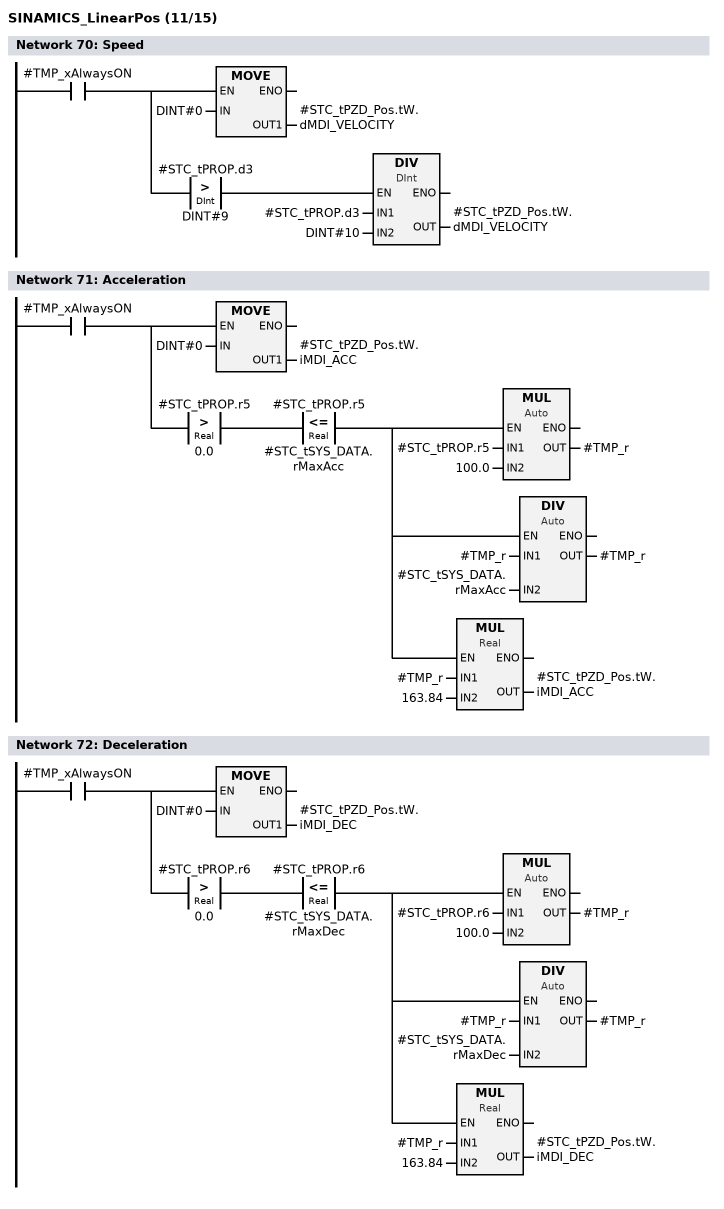
   RUNG wire#powerrail
      Contact( #TMP_xAlwaysON )
      wire#w1
      { S7_GenerateENO := "TRUE" } Move(in := DINT#0, out1 => #STC_tPZD_Pos.tW.dMDI_VELOCITY)
   END_RUNG
   RUNG wire#w1
      { S7_Templates := "SrcType := DInt" } GT_Contact(in1 := #STC_tPROP.d3, in2 := DINT#9)
      { S7_Templates := "SrcType := DInt"; S7_GenerateENO := "TRUE" } Div(in1 := #STC_tPROP.d3, in2 := DINT#10, out => #STC_tPZD_Pos.tW.dMDI_VELOCITY)
   END_RUNG
   // the same network as SCL:
   IF #TMP_xAlwaysON THEN #STC_tPZD_Pos.tW.dMDI_VELOCITY := DINT#0; END_IF;
   IF #TMP_xAlwaysON AND (#STC_tPROP.d3 > DINT#9) THEN
       #STC_tPZD_Pos.tW.dMDI_VELOCITY := #STC_tPROP.d3 / DINT#10;
   END_IF;
END_REGION

REGION Network 71: Acceleration
   RUNG wire#powerrail
      Contact( #TMP_xAlwaysON )
      wire#w1
      Move(in := DINT#0, out1 => #STC_tPZD_Pos.tW.iMDI_ACC)
   END_RUNG
   RUNG wire#w1
      { S7_Templates := "SrcType := Real" } GT_Contact(in1 := #STC_tPROP.r5, in2 := 0.0)
      { S7_Templates := "SrcType := Real" } LE_Contact(in1 := #STC_tPROP.r5, in2 := #STC_tSYS_DATA.rMaxAcc)
      wire#w2
      Mul(in1 := #STC_tPROP.r5, in2 := 100.0, out => #TMP_r)
   END_RUNG
   RUNG wire#w2
      Div(in1 := #TMP_r, in2 := #STC_tSYS_DATA.rMaxAcc, out => #TMP_r)
   END_RUNG
   RUNG wire#w2
      { S7_Templates := "SrcType := Real" } Mul(in1 := #TMP_r, in2 := 163.84, out => #STC_tPZD_Pos.tW.iMDI_ACC)
   END_RUNG
   // the same network as SCL:
   IF #TMP_xAlwaysON THEN #STC_tPZD_Pos.tW.iMDI_ACC := DINT#0; END_IF;
   IF #TMP_xAlwaysON AND (#STC_tPROP.r5 > 0.0) AND (#STC_tPROP.r5 <= #STC_tSYS_DATA.rMaxAcc) THEN
       #TMP_r := #STC_tPROP.r5 * 100.0;
       #TMP_r := #TMP_r / #STC_tSYS_DATA.rMaxAcc;
       #STC_tPZD_Pos.tW.iMDI_ACC := #TMP_r * 163.84;
   END_IF;
END_REGION

REGION Network 72: Deceleration
   RUNG wire#powerrail
      Contact( #TMP_xAlwaysON )
      wire#w1
      Move(in := DINT#0, out1 => #STC_tPZD_Pos.tW.iMDI_DEC)
   END_RUNG
   RUNG wire#w1
      { S7_Templates := "SrcType := Real" } GT_Contact(in1 := #STC_tPROP.r6, in2 := 0.0)
      { S7_Templates := "SrcType := Real" } LE_Contact(in1 := #STC_tPROP.r6, in2 := #STC_tSYS_DATA.rMaxDec)
      wire#w2
      Mul(in1 := #STC_tPROP.r6, in2 := 100.0, out => #TMP_r)
   END_RUNG
   RUNG wire#w2
      Div(in1 := #TMP_r, in2 := #STC_tSYS_DATA.rMaxDec, out => #TMP_r)
   END_RUNG
   RUNG wire#w2
      { S7_Templates := "SrcType := Real" } Mul(in1 := #TMP_r, in2 := 163.84, out => #STC_tPZD_Pos.tW.iMDI_DEC)
   END_RUNG
   // the same network as SCL:
   IF #TMP_xAlwaysON THEN #STC_tPZD_Pos.tW.iMDI_DEC := DINT#0; END_IF;
   IF #TMP_xAlwaysON AND (#STC_tPROP.r6 > 0.0) AND (#STC_tPROP.r6 <= #STC_tSYS_DATA.rMaxDec) THEN
       #TMP_r := #STC_tPROP.r6 * 100.0;
       #TMP_r := #TMP_r / #STC_tSYS_DATA.rMaxDec;
       #STC_tPZD_Pos.tW.iMDI_DEC := #TMP_r * 163.84;
   END_IF;
END_REGION

REGION Network 73: ########################_OPEN_CLOSE_LOOP_#######################
END_REGION

REGION Network 74: #####_MATCH_#####
END_REGION

REGION Network 75 (STL): Input copy
         JU    Out;

   T1:   CALL  BLKMOV
         ( SRCBLK  := #TMP_a,
           RET_VAL := #TMP_iRetVal,
           DSTBLK  := #STC_tPZD_OpCLLoop.tR
         );
END_REGION

REGION Network 76: Status signals
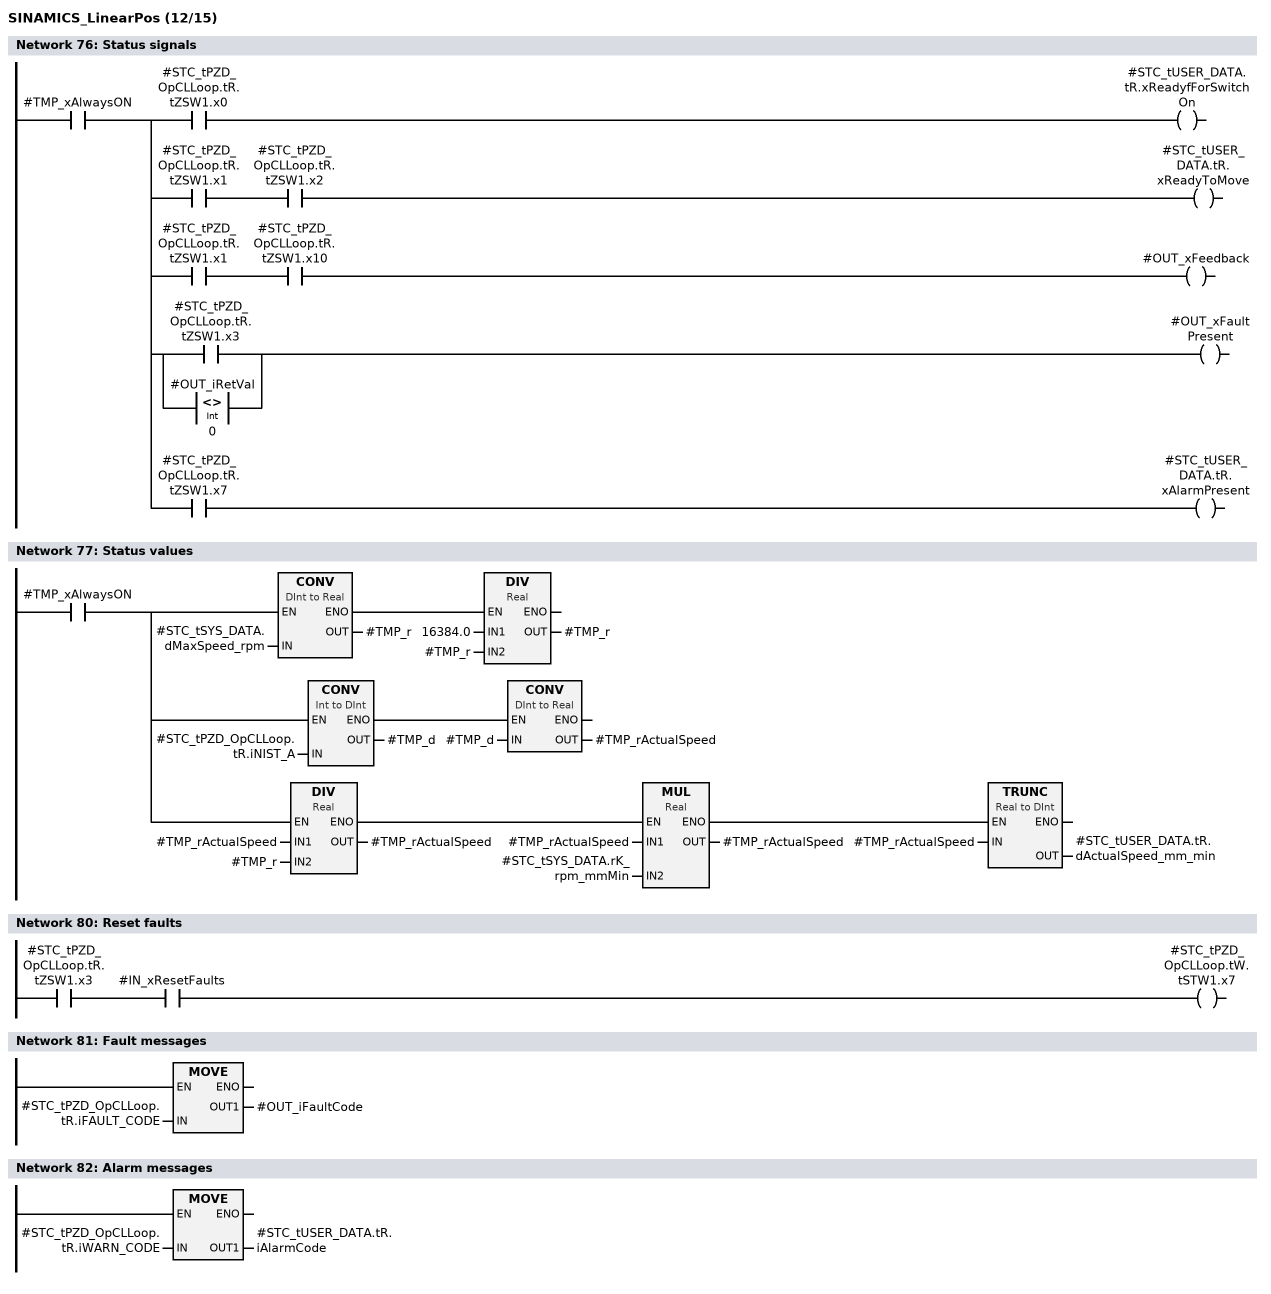
   RUNG wire#powerrail
      Contact( #TMP_xAlwaysON )
      wire#w1
      Contact( #STC_tPZD_OpCLLoop.tR.tZSW1.x0 )
      Coil( #STC_tUSER_DATA.tR.xReadyfForSwitchOn )
   END_RUNG
   RUNG wire#w1
      Contact( #STC_tPZD_OpCLLoop.tR.tZSW1.x1 )
      Contact( #STC_tPZD_OpCLLoop.tR.tZSW1.x2 )
      Coil( #STC_tUSER_DATA.tR.xReadyToMove )
   END_RUNG
   RUNG wire#w1
      Contact( #STC_tPZD_OpCLLoop.tR.tZSW1.x1 )
      Contact( #STC_tPZD_OpCLLoop.tR.tZSW1.x10 )
      Coil( #OUT_xFeedback )
   END_RUNG
   RUNG wire#w1
      Contact( #STC_tPZD_OpCLLoop.tR.tZSW1.x3 )
      wire#w2
      Coil( #OUT_xFaultPresent )
   END_RUNG
   RUNG wire#w1
      { S7_Templates := "SrcType := Int" } NE_Contact(in1 := #OUT_iRetVal, in2 := 0)
   END_RUNG wire#w2
   RUNG wire#w1
      Contact( #STC_tPZD_OpCLLoop.tR.tZSW1.x7 )
      Coil( #STC_tUSER_DATA.tR.xAlarmPresent )
   END_RUNG
   // the same network as SCL:
   #STC_tUSER_DATA.tR.xReadyfForSwitchOn := #TMP_xAlwaysON AND #STC_tPZD_OpCLLoop.tR.tZSW1.x0;
   #STC_tUSER_DATA.tR.xReadyToMove := #TMP_xAlwaysON AND #STC_tPZD_OpCLLoop.tR.tZSW1.x1 AND #STC_tPZD_OpCLLoop.tR.tZSW1.x2;
   #OUT_xFeedback := #TMP_xAlwaysON AND #STC_tPZD_OpCLLoop.tR.tZSW1.x1 AND #STC_tPZD_OpCLLoop.tR.tZSW1.x10;
   #OUT_xFaultPresent := #TMP_xAlwaysON AND (#STC_tPZD_OpCLLoop.tR.tZSW1.x3 OR (#OUT_iRetVal <> 0));
   #STC_tUSER_DATA.tR.xAlarmPresent := #TMP_xAlwaysON AND #STC_tPZD_OpCLLoop.tR.tZSW1.x7;
END_REGION

REGION Network 77: Status values
   RUNG wire#powerrail
      Contact( #TMP_xAlwaysON )
      wire#w1
      { S7_Templates := "[SrcType := DInt, DestType := Real]"; S7_GenerateENO := "TRUE" } Convert(in := #STC_tSYS_DATA.dMaxSpeed_rpm, out => #TMP_r)
      { S7_Templates := "SrcType := Real"; S7_GenerateENO := "TRUE" } Div(in1 := 16384.0, in2 := #TMP_r, out => #TMP_r)
   END_RUNG
   RUNG wire#w1
      { S7_Templates := "[SrcType := Int, DestType := DInt]"; S7_GenerateENO := "TRUE" } Convert(in := #STC_tPZD_OpCLLoop.tR.iNIST_A, out => #TMP_d)
      { S7_Templates := "[SrcType := DInt, DestType := Real]"; S7_GenerateENO := "TRUE" } Convert(in := #TMP_d, out => #TMP_rActualSpeed)
   END_RUNG
   RUNG wire#w1
      { S7_Templates := "SrcType := Real"; S7_GenerateENO := "TRUE" } Div(in1 := #TMP_rActualSpeed, in2 := #TMP_r, out => #TMP_rActualSpeed)
      { S7_Templates := "SrcType := Real"; S7_GenerateENO := "TRUE" } Mul(in1 := #TMP_rActualSpeed, in2 := #STC_tSYS_DATA.rK_rpm_mmMin, out => #TMP_rActualSpeed)
      { S7_Templates := "[SrcType := Real, DestType := DInt]"; S7_GenerateENO := "TRUE" } Trunc(in := #TMP_rActualSpeed, out => #STC_tUSER_DATA.tR.dActualSpeed_mm_min)
   END_RUNG
   // the same network as SCL:
   // ENO of a box is taken as its EN; it also drops when the box reports an error
   IF #TMP_xAlwaysON THEN
       #TMP_r := DINT_TO_REAL(#STC_tSYS_DATA.dMaxSpeed_rpm);
       #TMP_r := 16384.0 / #TMP_r;
       #TMP_d := INT_TO_DINT(#STC_tPZD_OpCLLoop.tR.iNIST_A);
       #TMP_rActualSpeed := DINT_TO_REAL(#TMP_d);
       #TMP_rActualSpeed := #TMP_rActualSpeed / #TMP_r;
       #TMP_rActualSpeed := #TMP_rActualSpeed * #STC_tSYS_DATA.rK_rpm_mmMin;
       #STC_tUSER_DATA.tR.dActualSpeed_mm_min := TRUNC(#TMP_rActualSpeed);
   END_IF;
END_REGION

REGION Network 78: #####_STATUSES_#####
END_REGION

REGION Network 79: #####_ALARMS_#####
END_REGION

REGION Network 80: Reset faults
   RUNG wire#powerrail
      Contact( #STC_tPZD_OpCLLoop.tR.tZSW1.x3 )
      Contact( #IN_xResetFaults )
      Coil( #STC_tPZD_OpCLLoop.tW.tSTW1.x7 )
   END_RUNG
   // the same network as SCL:
   #STC_tPZD_OpCLLoop.tW.tSTW1.x7 := #STC_tPZD_OpCLLoop.tR.tZSW1.x3 AND #IN_xResetFaults;
END_REGION

REGION Network 81: Fault messages
   RUNG wire#powerrail
      { S7_GenerateENO := "TRUE" } Move(in := #STC_tPZD_OpCLLoop.tR.iFAULT_CODE, out1 => #OUT_iFaultCode)
   END_RUNG
   // the same network as SCL:
   #OUT_iFaultCode := #STC_tPZD_OpCLLoop.tR.iFAULT_CODE;
END_REGION

REGION Network 82: Alarm messages
   RUNG wire#powerrail
      { S7_GenerateENO := "TRUE" } Move(in := #STC_tPZD_OpCLLoop.tR.iWARN_CODE, out1 => #STC_tUSER_DATA.tR.iAlarmCode)
   END_RUNG
   // the same network as SCL:
   #STC_tUSER_DATA.tR.iAlarmCode := #STC_tPZD_OpCLLoop.tR.iWARN_CODE;
END_REGION

REGION Network 83: #####_PHASES_&_LOGICS_#####
END_REGION

REGION Network 84: Enable PLC control
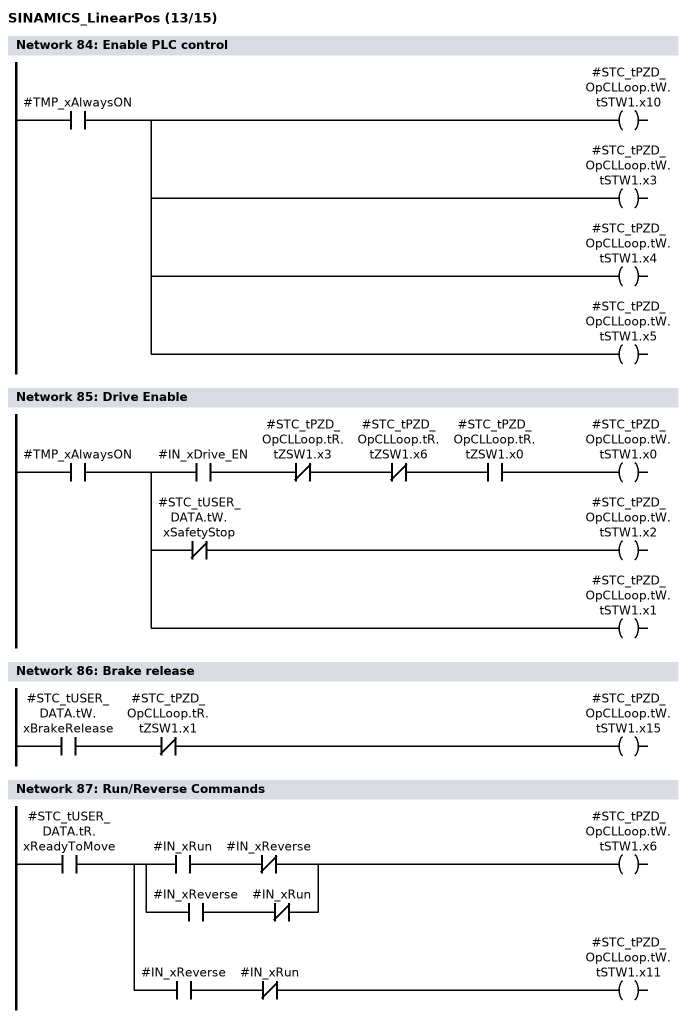
   RUNG wire#powerrail
      Contact( #TMP_xAlwaysON )
      wire#w1
      Coil( #STC_tPZD_OpCLLoop.tW.tSTW1.x10 )
   END_RUNG
   RUNG wire#w1
      Coil( #STC_tPZD_OpCLLoop.tW.tSTW1.x3 )
   END_RUNG
   RUNG wire#w1
      Coil( #STC_tPZD_OpCLLoop.tW.tSTW1.x4 )
   END_RUNG
   RUNG wire#w1
      Coil( #STC_tPZD_OpCLLoop.tW.tSTW1.x5 )
   END_RUNG
   // the same network as SCL:
   #STC_tPZD_OpCLLoop.tW.tSTW1.x10 := #TMP_xAlwaysON;
   #STC_tPZD_OpCLLoop.tW.tSTW1.x3 := #TMP_xAlwaysON;
   #STC_tPZD_OpCLLoop.tW.tSTW1.x4 := #TMP_xAlwaysON;
   #STC_tPZD_OpCLLoop.tW.tSTW1.x5 := #TMP_xAlwaysON;
END_REGION

REGION Network 85: Drive Enable
   RUNG wire#powerrail
      Contact( #TMP_xAlwaysON )
      wire#w1
      Contact( #IN_xDrive_EN )
      I_Contact( #STC_tPZD_OpCLLoop.tR.tZSW1.x3 )
      I_Contact( #STC_tPZD_OpCLLoop.tR.tZSW1.x6 )
      Contact( #STC_tPZD_OpCLLoop.tR.tZSW1.x0 )
      Coil( #STC_tPZD_OpCLLoop.tW.tSTW1.x0 )
   END_RUNG
   RUNG wire#w1
      I_Contact( #STC_tUSER_DATA.tW.xSafetyStop )
      Coil( #STC_tPZD_OpCLLoop.tW.tSTW1.x2 )
   END_RUNG
   RUNG wire#w1
      Coil( #STC_tPZD_OpCLLoop.tW.tSTW1.x1 )
   END_RUNG
   // the same network as SCL:
   #STC_tPZD_OpCLLoop.tW.tSTW1.x0 := #TMP_xAlwaysON AND #IN_xDrive_EN AND NOT #STC_tPZD_OpCLLoop.tR.tZSW1.x3 AND NOT #STC_tPZD_OpCLLoop.tR.tZSW1.x6 AND #STC_tPZD_OpCLLoop.tR.tZSW1.x0;
   #STC_tPZD_OpCLLoop.tW.tSTW1.x2 := #TMP_xAlwaysON AND NOT #STC_tUSER_DATA.tW.xSafetyStop;
   #STC_tPZD_OpCLLoop.tW.tSTW1.x1 := #TMP_xAlwaysON;
END_REGION

REGION Network 86: Brake release
   RUNG wire#powerrail
      Contact( #STC_tUSER_DATA.tW.xBrakeRelease )
      I_Contact( #STC_tPZD_OpCLLoop.tR.tZSW1.x1 )
      Coil( #STC_tPZD_OpCLLoop.tW.tSTW1.x15 )
   END_RUNG
   // the same network as SCL:
   #STC_tPZD_OpCLLoop.tW.tSTW1.x15 := #STC_tUSER_DATA.tW.xBrakeRelease AND NOT #STC_tPZD_OpCLLoop.tR.tZSW1.x1;
END_REGION

REGION Network 87: Run/Reverse Commands
   RUNG wire#powerrail
      Contact( #STC_tUSER_DATA.tR.xReadyToMove )
      wire#w1
      Contact( #IN_xRun )
      I_Contact( #IN_xReverse )
      wire#w2
      Coil( #STC_tPZD_OpCLLoop.tW.tSTW1.x6 )
   END_RUNG
   RUNG wire#w1
      Contact( #IN_xReverse )
      I_Contact( #IN_xRun )
   END_RUNG wire#w2
   RUNG wire#w1
      Contact( #IN_xReverse )
      I_Contact( #IN_xRun )
      Coil( #STC_tPZD_OpCLLoop.tW.tSTW1.x11 )
   END_RUNG
   // the same network as SCL:
   #STC_tPZD_OpCLLoop.tW.tSTW1.x6 := #STC_tUSER_DATA.tR.xReadyToMove AND ((#IN_xRun AND NOT #IN_xReverse) OR (#IN_xReverse AND NOT #IN_xRun));
   #STC_tPZD_OpCLLoop.tW.tSTW1.x11 := #STC_tUSER_DATA.tR.xReadyToMove AND #IN_xReverse AND NOT #IN_xRun;
END_REGION

REGION Network 88: #####_PARAMETERS_#####
END_REGION

REGION Network 89: Speed
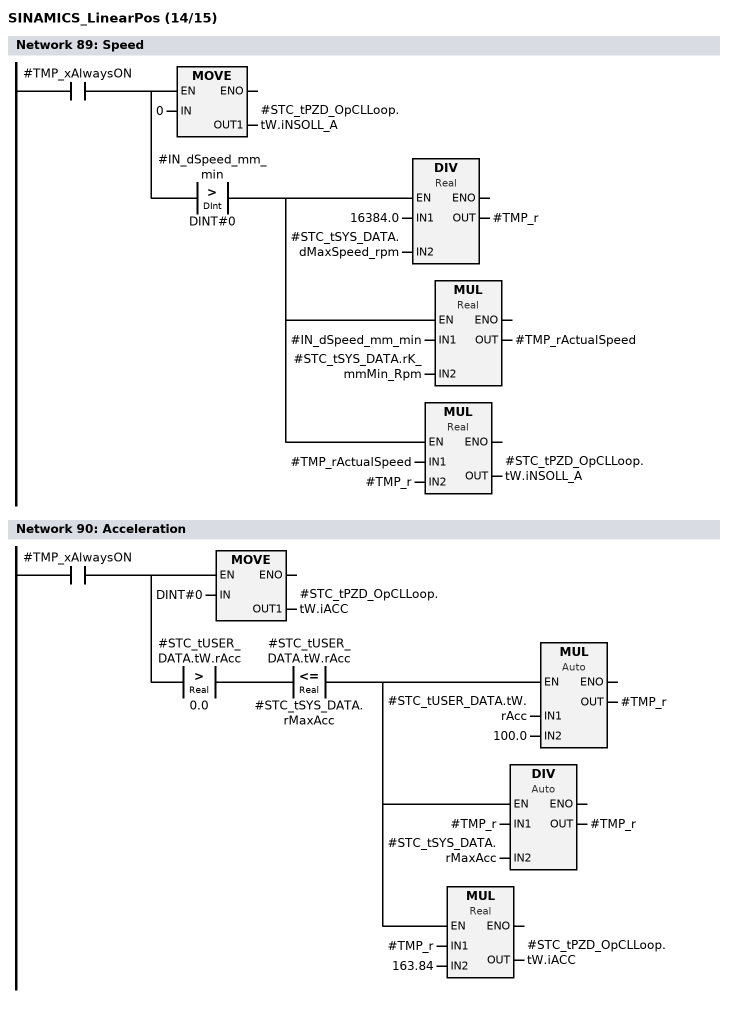
   RUNG wire#powerrail
      Contact( #TMP_xAlwaysON )
      wire#w1
      Move(in := 0, out1 => #STC_tPZD_OpCLLoop.tW.iNSOLL_A)
   END_RUNG
   RUNG wire#w1
      { S7_Templates := "SrcType := DInt" } GT_Contact(in1 := #IN_dSpeed_mm_min, in2 := DINT#0)
      wire#w2
      { S7_Templates := "SrcType := Real" } Div(in1 := 16384.0, in2 := #STC_tSYS_DATA.dMaxSpeed_rpm, out => #TMP_r)
   END_RUNG
   RUNG wire#w2
      { S7_Templates := "SrcType := Real" } Mul(in1 := #IN_dSpeed_mm_min, in2 := #STC_tSYS_DATA.rK_mmMin_Rpm, out => #TMP_rActualSpeed)
   END_RUNG
   RUNG wire#w2
      { S7_Templates := "SrcType := Real" } Mul(in1 := #TMP_rActualSpeed, in2 := #TMP_r, out => #STC_tPZD_OpCLLoop.tW.iNSOLL_A)
   END_RUNG
   // the same network as SCL:
   IF #TMP_xAlwaysON THEN #STC_tPZD_OpCLLoop.tW.iNSOLL_A := 0; END_IF;
   IF #TMP_xAlwaysON AND (#IN_dSpeed_mm_min > DINT#0) THEN
       #TMP_r := 16384.0 / #STC_tSYS_DATA.dMaxSpeed_rpm;
       #TMP_rActualSpeed := #IN_dSpeed_mm_min * #STC_tSYS_DATA.rK_mmMin_Rpm;
       #STC_tPZD_OpCLLoop.tW.iNSOLL_A := #TMP_rActualSpeed * #TMP_r;
   END_IF;
END_REGION

REGION Network 90: Acceleration
   RUNG wire#powerrail
      Contact( #TMP_xAlwaysON )
      wire#w1
      Move(in := DINT#0, out1 => #STC_tPZD_OpCLLoop.tW.iACC)
   END_RUNG
   RUNG wire#w1
      { S7_Templates := "SrcType := Real" } GT_Contact(in1 := #STC_tUSER_DATA.tW.rAcc, in2 := 0.0)
      { S7_Templates := "SrcType := Real" } LE_Contact(in1 := #STC_tUSER_DATA.tW.rAcc, in2 := #STC_tSYS_DATA.rMaxAcc)
      wire#w2
      Mul(in1 := #STC_tUSER_DATA.tW.rAcc, in2 := 100.0, out => #TMP_r)
   END_RUNG
   RUNG wire#w2
      Div(in1 := #TMP_r, in2 := #STC_tSYS_DATA.rMaxAcc, out => #TMP_r)
   END_RUNG
   RUNG wire#w2
      { S7_Templates := "SrcType := Real" } Mul(in1 := #TMP_r, in2 := 163.84, out => #STC_tPZD_OpCLLoop.tW.iACC)
   END_RUNG
   // the same network as SCL:
   IF #TMP_xAlwaysON THEN #STC_tPZD_OpCLLoop.tW.iACC := DINT#0; END_IF;
   IF #TMP_xAlwaysON AND (#STC_tUSER_DATA.tW.rAcc > 0.0) AND (#STC_tUSER_DATA.tW.rAcc <= #STC_tSYS_DATA.rMaxAcc) THEN
       #TMP_r := #STC_tUSER_DATA.tW.rAcc * 100.0;
       #TMP_r := #TMP_r / #STC_tSYS_DATA.rMaxAcc;
       #STC_tPZD_OpCLLoop.tW.iACC := #TMP_r * 163.84;
   END_IF;
END_REGION

REGION Network 91: Deceleration
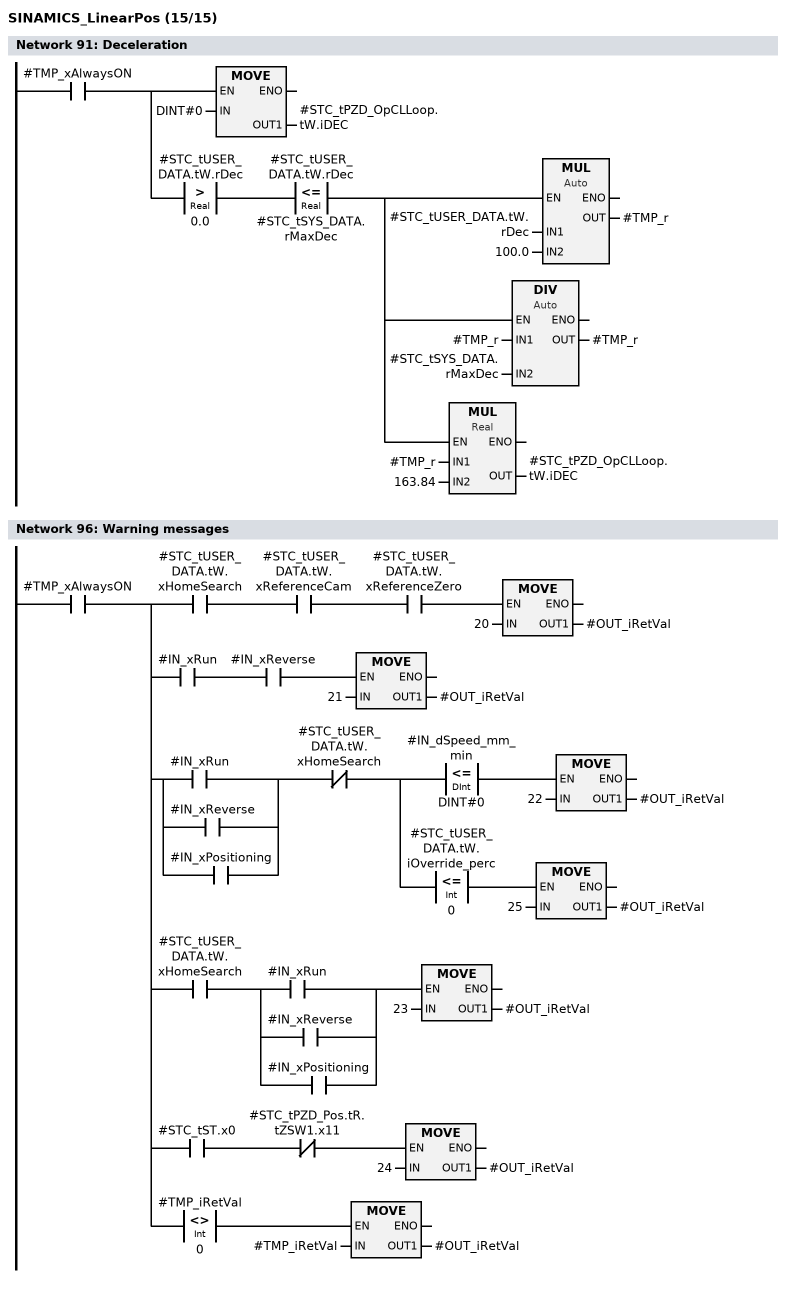
   RUNG wire#powerrail
      Contact( #TMP_xAlwaysON )
      wire#w1
      Move(in := DINT#0, out1 => #STC_tPZD_OpCLLoop.tW.iDEC)
   END_RUNG
   RUNG wire#w1
      { S7_Templates := "SrcType := Real" } GT_Contact(in1 := #STC_tUSER_DATA.tW.rDec, in2 := 0.0)
      { S7_Templates := "SrcType := Real" } LE_Contact(in1 := #STC_tUSER_DATA.tW.rDec, in2 := #STC_tSYS_DATA.rMaxDec)
      wire#w2
      Mul(in1 := #STC_tUSER_DATA.tW.rDec, in2 := 100.0, out => #TMP_r)
   END_RUNG
   RUNG wire#w2
      Div(in1 := #TMP_r, in2 := #STC_tSYS_DATA.rMaxDec, out => #TMP_r)
   END_RUNG
   RUNG wire#w2
      { S7_Templates := "SrcType := Real" } Mul(in1 := #TMP_r, in2 := 163.84, out => #STC_tPZD_OpCLLoop.tW.iDEC)
   END_RUNG
   // the same network as SCL:
   IF #TMP_xAlwaysON THEN #STC_tPZD_OpCLLoop.tW.iDEC := DINT#0; END_IF;
   IF #TMP_xAlwaysON AND (#STC_tUSER_DATA.tW.rDec > 0.0) AND (#STC_tUSER_DATA.tW.rDec <= #STC_tSYS_DATA.rMaxDec) THEN
       #TMP_r := #STC_tUSER_DATA.tW.rDec * 100.0;
       #TMP_r := #TMP_r / #STC_tSYS_DATA.rMaxDec;
       #STC_tPZD_OpCLLoop.tW.iDEC := #TMP_r * 163.84;
   END_IF;
END_REGION

REGION Network 92: ################_MOTOR_MODULE_TELEGRAMS_ENDING_#################
END_REGION

REGION Network 93 (STL): Output copy motor module
   Out:  L     #STC_tSYS_DATA.iPZD_MM;
         L     111;
         ==I;
         L     12;
         T     #TMP_iAddressLength;
         JC    WOut;
         L     #STC_tSYS_DATA.iPZD_MM;
         L     1;
         ==I;
         L     4;
         T     #TMP_iAddressLength;
         JC    WOut;

         L     19;
         JU    Err;

   WOut: NOP   0;

   //Compute destination position
         L;
         LAR1;
   //byte 1 = 10h (FIXED for S7)
         L     B#16#10;
         T     B[AR1, P#0.0];
   //byte 2 = data type
         L     B#16#4;  //4 = word
         T     B[AR1, P#1.0];
   //byte 3 & 4 = number of element
         L     #TMP_iAddressLength;  //Production data
         T     W[AR1, P#2.0];
   //byte 5 & 6 = number of DB
         L     0;  //DB production data
         T     W[AR1, P#4.0];
   //byte 7 = memory area
         L     B#16#82;  //82h = Q (Output)
         T     B[AR1, P#6.0];
   //byte 8 & 9 = address. Bit 0,1,2 of tenth byte is bit offset
   //byte 7 = address (high). Valid value = 0-7. Bit 3,4,5,6,7 always 0
         L     #STC_tSYS_DATA.iIOAddress_MM;  //Item size
         SLW   3;
         T     W[AR1, P#8.0];
         SRD   16;
         AW    16#0007;
         T     B[AR1, P#7.0];

         L     #STC_tSYS_DATA.iPZD_MM;
         L     1;
         ==I;
         JC    W1;

         CALL  BLKMOV
         ( SRCBLK  := #STC_tPZD_Pos.tW,
           RET_VAL := #TMP_iRetVal,
           DSTBLK  := #TMP_a
         );

         JU    WEnd;

   W1:   CALL  BLKMOV
         ( SRCBLK  := #STC_tPZD_OpCLLoop.tW,
           RET_VAL := #TMP_iRetVal,
           DSTBLK  := #TMP_a
         );

   WEnd: NOP   0;
END_REGION

REGION Network 94: #####_RETVAL_RESPONSE_#####
END_REGION

REGION Network 95 (STL): Initialize RetVal
         L     0;
         T     #OUT_iRetVal;
END_REGION

REGION Network 96: Warning messages
   RUNG wire#powerrail
      Contact( #TMP_xAlwaysON )
      wire#w1
      Contact( #STC_tUSER_DATA.tW.xHomeSearch )
      Contact( #STC_tUSER_DATA.tW.xReferenceCam )
      Contact( #STC_tUSER_DATA.tW.xReferenceZero )
      Move(in := 20, out1 => #OUT_iRetVal)
   END_RUNG
   RUNG wire#w1
      Contact( #IN_xRun )
      Contact( #IN_xReverse )
      Move(in := 21, out1 => #OUT_iRetVal)
   END_RUNG
   RUNG wire#w1
      Contact( #IN_xRun )
      wire#w2
      I_Contact( #STC_tUSER_DATA.tW.xHomeSearch )
      wire#w3
      { S7_Templates := "SrcType := DInt" } LE_Contact(in1 := #IN_dSpeed_mm_min, in2 := DINT#0)
      Move(in := 22, out1 => #OUT_iRetVal)
   END_RUNG
   RUNG wire#w1
      Contact( #IN_xReverse )
   END_RUNG wire#w2
   RUNG wire#w1
      Contact( #IN_xPositioning )
   END_RUNG wire#w2
   RUNG wire#w3
      { S7_Templates := "SrcType := Int" } LE_Contact(in1 := #STC_tUSER_DATA.tW.iOverride_perc, in2 := 0)
      Move(in := 25, out1 => #OUT_iRetVal)
   END_RUNG
   RUNG wire#w1
      Contact( #STC_tUSER_DATA.tW.xHomeSearch )
      wire#w4
      Contact( #IN_xRun )
      wire#w5
      Move(in := 23, out1 => #OUT_iRetVal)
   END_RUNG
   RUNG wire#w4
      Contact( #IN_xReverse )
   END_RUNG wire#w5
   RUNG wire#w4
      Contact( #IN_xPositioning )
   END_RUNG wire#w5
   RUNG wire#w1
      Contact( #STC_tST.x0 )
      I_Contact( #STC_tPZD_Pos.tR.tZSW1.x11 )
      Move(in := 24, out1 => #OUT_iRetVal)
   END_RUNG
   RUNG wire#w1
      { S7_Templates := "SrcType := Int" } NE_Contact(in1 := #TMP_iRetVal, in2 := 0)
      Move(in := #TMP_iRetVal, out1 => #OUT_iRetVal)
   END_RUNG
   // the same network as SCL:
   IF #TMP_xAlwaysON AND #STC_tUSER_DATA.tW.xHomeSearch AND #STC_tUSER_DATA.tW.xReferenceCam AND #STC_tUSER_DATA.tW.xReferenceZero THEN
       #OUT_iRetVal := 20;
   END_IF;
   IF #TMP_xAlwaysON AND #IN_xRun AND #IN_xReverse THEN #OUT_iRetVal := 21; END_IF;
   #_w1 := #TMP_xAlwaysON AND (#IN_xRun OR #IN_xReverse OR #IN_xPositioning) AND NOT #STC_tUSER_DATA.tW.xHomeSearch;
   IF #_w1 AND (#IN_dSpeed_mm_min <= DINT#0) THEN #OUT_iRetVal := 22; END_IF;
   IF #_w1 AND (#STC_tUSER_DATA.tW.iOverride_perc <= 0) THEN #OUT_iRetVal := 25; END_IF;
   IF #TMP_xAlwaysON AND #STC_tUSER_DATA.tW.xHomeSearch AND (#IN_xRun OR #IN_xReverse OR #IN_xPositioning) THEN
       #OUT_iRetVal := 23;
   END_IF;
   IF #TMP_xAlwaysON AND #STC_tST.x0 AND NOT #STC_tPZD_Pos.tR.tZSW1.x11 THEN #OUT_iRetVal := 24; END_IF;
   IF #TMP_xAlwaysON AND (#TMP_iRetVal <> 0) THEN #OUT_iRetVal := #TMP_iRetVal; END_IF;
END_REGION

REGION Network 97 (STL): Blocking messages
         JU    Rest;
   Err:  T     #OUT_iRetVal;
END_REGION

REGION Network 98 (STL): Reset input commands
   // R     #USER_DATA.W.SafetyStop
   //       R     #USER_DATA.W.FlyChange
   //       R     #USER_DATA.W.PH_Select
   //       R     #USER_DATA.W.StartCountOnHead
   //       R     #USER_DATA.W.StartCountOnTail
   //       R     #USER_DATA.W.BrakeRelease
   //       R     #USER_DATA.W.ResetCount
   //       R     #USER_DATA.W.PresetRq
   //       R     #USER_DATA.W.HomeSearch
   //       R     #USER_DATA.W.ReverseHoming
   //       R     #USER_DATA.W.ReferenceCam
   //       R     #USER_DATA.W.ReferenceZero
   //       R     #USER_DATA.W.MDI_Continue
   //       R     #USER_DATA.W.SwLimitsEnable
   //       R     #USER_DATA.W.HwLimitsEnable
   //       R     #Run
   //       R     #Reverse
   //       R     #Positioning
   // 
   //       L     L#0
   //       T     #Speed
   //       T     #USER_DATA.W.Override
   //       T     #USER_DATA.W.Target
   //       T     #USER_DATA.W.Preset
   //       T     #USER_DATA.W.Acc
   //       T     #USER_DATA.W.Dec
   Rest: NOP   0;
   //    SET
   //    R     #IN_xDrive_EN
   //    R     #IN_xResetFaults
END_REGION

REGION Network 99 (STL): Restore AR1 & AR2 value
   //    L     #TMP_dOldValue_AR1
   //    LAR1
   //    L     #TMP_dOldValue_AR2
   //    LAR2
END_REGION
END_FUNCTION_BLOCK

FUNCTION_BLOCK "SINAMICS_RotativePos"   // FB52, LAD
TITLE = Sinamics drive manager
{ S7_Optimized_Access := 'FALSE' }
AUTHOR : Armitano
VERSION : 1.4
   VAR_INPUT
      IN_xDrive_EN : Bool;   // Drive enable
      IN_xRun : Bool;   // Run clockwise
      IN_xReverse : Bool;   // Run counterclockwise
      IN_xPositioning : Bool;   // Positioning enable
      IN_xResetFaults : Bool;   // Reset faults
      IN_dSpeed_deg_min : DInt;   // Speed reference [°/min]
   END_VAR
   VAR_OUTPUT
      OUT_xFeedback : Bool;   // Feedback active
      OUT_xFaultPresent : Bool;   // Fault present
      OUT_iFaultCode : Int;   // Fault code
      OUT_iRetVal : Int;   // Return value in case of wrong configuration
   END_VAR
   VAR
      STC_tUSER_DATA : Struct   // User data (Extended functions commands for execute the application desired)
         tR : Struct
            xReadyfForSwitchOn : Bool;   // Ready for switch on
            xReadyToMove : Bool;   // Ready to move
            xAxleRefered : Bool;   // Axle referenced
            xPositionReached : Bool;   // Position reached
            xAlarmPresent : Bool;   // Alarm present
            xAxleToZero : Bool;   // Axle to zero value (only positioner)
            iAlarmCode : Int;   // Alarm code
            dActualPosition_cdeg : DInt;   // Actual position value [°/100]
            dActualSpeed_deg_min : DInt;   // Actual speed value [°/min]
         END_STRUCT;
         tW : Struct
            xSafetyStop : Bool;   // Safety stop (OFF3)
            xFlyChange : Bool;   // Fly change
            x3 : Bool;
            x4 : Bool;
            x5 : Bool;
            xBrakeRelease : Bool;   // Brake release
            xResetCount : Bool;   // Reset counter
            xPresetRq : Bool;   // Preset request (only absolute encoder)
            xHomeSearch : Bool;   // Home search cycle (only for homing)
            xReverseHoming : Bool;   // Reverse homing search direction (only for homing)
            xReferenceCam : Bool;   // Sensor reference cam for homing cycle + zero mark (only for homing)
            xReferenceZero : Bool;   // Sensor reference zero for homing cycle (only for homing)
            xMDI_Continue : Bool;   // MDI movment continue (only for gearing axes)
            x14 : Bool;
            xHwLimitsEnable : Bool;   // Hardware limits activation (only positioner)
            iOverride_perc : Int := 100;   // Override [%]
            dTarget_cdeg : DInt;   // Target position [°/100]
            dPreset_cdeg : DInt;   // Preset position [°/100] (only for homing & absolute encoder)
            rAcc_deg_s2 : Real;   // Acceleration [°/s2]
            rDec_deg_s2 : Real;   // Deceleration [°/s2]
         END_STRUCT;
      END_STRUCT;
      STC_tSYS_DATA : Struct   // System data (Info about applications type and HW config.)
         iIOAddress_MM : Int := -1;   // Input/Output addresses for motor module
         i2 : Int;
         i3 : Int;
         iDiagAddress : Int;   // Diagnostic address of SINAMICS module (only for absolute encoder & homing)
         iPosPZD_CU : Int;   // Number of PZD position in SINAMICS configuration [1,2,3..] (for absolute enc.)
         iPosPZD_MM : Int;   // Number of PZD position in SINAMICS configuration [1,2,3..] (for homing & enc.)
         i7 : Int;
         dMaxSpeed_rpm : DInt;   // MaxSpeed [rpm]
         d9 : DInt;
         dPosWindow_cdeg : DInt := L#40;   // Positioning window [°/100]
         d11 : DInt;
         d12 : DInt;
         d13 : DInt;
         rK_rpm_degMin : Real;   // K Conversion from rpm to °/min
         r15 : Real;
         rMaxAcc_deg_s2 : Real;   // MaxAcc [°/s2]
         rMaxDec_deg_s2 : Real;   // MaxDec [°/s2]
         r18 : Real;
         r19 : Real;
      END_STRUCT;
      STC_tEXT_DATA : Struct   // Extended data (Special functions commands for extra applications)
         tR : Struct
            x0 : Bool;
            x1 : Bool;
            x2 : Bool;
            x3 : Bool;
            x4 : Bool;
            x5 : Bool;
            x6 : Bool;
            x7 : Bool;
            x8 : Bool;
            x9 : Bool;
            x10 : Bool;
            x11 : Bool;
            x12 : Bool;
            x13 : Bool;
            x14 : Bool;
            x15 : Bool;
            d0 : DInt;
            d1 : DInt;
            d2 : DInt;
            d3 : DInt;
            d4 : DInt;
            d5 : DInt;
            d6 : DInt;
            d7 : DInt;
            d8 : DInt;
            d9 : DInt;
            d10 : DInt;
            d11 : DInt;
            rgdSpare : Array[0..5] of DInt;
         END_STRUCT;
         tW : Struct
            xDisGearingCtrl : Bool;   // Disable gearing tollerance error control (Only for gearing axes)
            x1 : Bool;
            x2 : Bool;
            x3 : Bool;
            x4 : Bool;
            xModuleCorrect : Bool;   // Enable module correction (only positioner with turnover endless)
            x6 : Bool;
            x7 : Bool;
            x8 : Bool;
            x9 : Bool;
            x10 : Bool;
            x11 : Bool;
            x12 : Bool;
            x13 : Bool;
            x14 : Bool;
            x15 : Bool;
            d0 : DInt;
            d1 : DInt;
            d2 : DInt;
            d3 : DInt;
            d4 : DInt;
            d5 : DInt;
            d6 : DInt;
            d7 : DInt;
            d8 : DInt;
            d9 : DInt;
            d10 : DInt;
            d11 : DInt;
            rgdSpare : Array[0..5] of DInt;
         END_STRUCT;
      END_STRUCT;
      STC_tST : Struct
         x0 : Bool;
         x1 : Bool;
         x2 : Bool;
         x3 : Bool;
         x4 : Bool;
         x5 : Bool;
         x6 : Bool;   // Target = Feedback target
         x7 : Bool;
         x8 : Bool;   // Preset phases in progress
         x9 : Bool;
         x10 : Bool;
         x11 : Bool;   // Axle resetted
         x12 : Bool;
         x13 : Bool;
         x14 : Bool;
         x15 : Bool;
      END_STRUCT;
      STC_tOS_PN : Struct
         x0 : Bool;   // Run
         x1 : Bool;   // Reverse
         x2 : Bool;   // Positioning
         x3 : Bool;   // Fly change
         x4 : Bool;
         x5 : Bool;
         x6 : Bool;
         x7 : Bool;
         x8 : Bool;
         x9 : Bool;
         x10 : Bool;   // Preset position
         x11 : Bool;
         x12 : Bool;
         x13 : Bool;
         x14 : Bool;
         x15 : Bool;
      END_STRUCT;
      STC_tOS : Struct
         x0 : Bool;   // Run
         x1 : Bool;   // Reverse
         x2 : Bool;   // Positioning
         x3 : Bool;   // Fly change
         x4 : Bool;
         x5 : Bool;
         x6 : Bool;
         x7 : Bool;
         x8 : Bool;
         x9 : Bool;
         x10 : Bool;
         x11 : Bool;
         x12 : Bool;
         x13 : Bool;
         x14 : Bool;
         x15 : Bool;
      END_STRUCT;
      STC_tPH : Struct
         x0 : Bool;   // Positioning initializing
         x1 : Bool;   // Positioning request
         x2 : Bool;   // Fly change waiting
         x3 : Bool;   // Fly change sending
         x4 : Bool;   // Change command waiting
         x5 : Bool;   // Change command request
         x6 : Bool;
         x7 : Bool;
         x8 : Bool;   // Send encoder value
         x9 : Bool;
         x10 : Bool;   // Send preset command
         x11 : Bool;
         x12 : Bool;   // Send saving preset command
         x13 : Bool;
         x14 : Bool;   // End preset encoder
         x15 : Bool;
      END_STRUCT;
      STC_tPROP : Struct
         i0 : Int;   // Previous cycle [ms]
         i1 : Int;
         i2 : Int;   // Override in sending [%]
         d3 : DInt;   // Speed in sending [°/min]
         d4 : DInt;   // Target in sending [°/100]
         r5 : Real;   // Acceleration in sending [°/s2]
         r6 : Real;   // Deceleration in sending [°/s2]
         i7 : Int;
         i8 : Int;
         i9 : Int;
         i10 : Int;
         i11 : Int;   // Override in fly change [%]
         d12 : DInt;   // Speed in fly change [°/min]
         d13 : DInt;   // Target in fly change [°/100]
         r14 : Real;   // Acceleration in fly change [°/s2]
         r15 : Real;   // Deceleration in fly change [°/s2]
         i16 : Int;
         i17 : Int;
         i18 : Int;
         i19 : Int;
         i20 : Int;
         tmON_feedback_ms : IEC_TIMER;   // Delay feedback [ms]
      END_STRUCT;
      STC_tR_MngSysReg : Struct   // Managment system register
         tST : Struct
            xRead_Request : Bool;
            xDone : Bool;
            xBusy : Bool;
            xError : Bool;
            xSpare4 : Bool;
            xSpare5 : Bool;
            xSpare6 : Bool;
            xSpare7 : Bool;
            ID : Hw_Io;
            dINDEX : DInt;
            uiLEN : UInt;
            dwSTATUS : DWord;
            uiMLEN : UInt;
         END_STRUCT;
         tDATA : Struct
            tRequestValues : Struct
               wRequest_refere_RequestID : Word := W#16#501;   // (Request_referece=01 Alwais=01 )*(RequestID=01 Read Param)
               wAxis_NoOfParameters : Word := W#16#112;   // (Axis=Num.Object)(NoOfParameters=Num of parameter to Read)
               wAttribute_NoOfElements_1 : Word := W#16#1000;   // (Attribute=10 Alwais=10)(NoOfParameters=Num of subparameter to Read)
               iParameter_number_1 : Int := 21700;   // Parameter_number=Number of the parameter
               wSubindex_1 : Word;   // Subindex
               wAttribute_NoOfElements_2 : Word := W#16#1000;   // (Attribute=10 Alwais=10)(NoOfParameters=Num of subparameter to Read)
               iParameter_number_2 : Int := 21701;   // Parameter_number=Number of the parameter
               wSubindex_2 : Word;   // Subindex
               wAttribute_NoOfElements_3 : Word := W#16#1000;   // (Attribute=10 Alwais=10)(NoOfParameters=Num of subparameter to Read)
               iParameter_number_3 : Int := 21702;   // Parameter_number=Number of the parameter
               wSubindex_3 : Word;   // Subindex
               wAttribute_NoOfElements_4 : Word := W#16#1000;   // (Attribute=10 Alwais=10)(NoOfParameters=Num of subparameter to Read)
               iParameter_number_4 : Int := 21703;   // Parameter_number=Number of the parameter
               wSubindex_4 : Word;   // Subindex
               wAttribute_NoOfElements_5 : Word := W#16#1000;   // (Attribute=10 Alwais=10)(NoOfParameters=Num of subparameter to Read)
               iParameter_number_5 : Int := 21704;   // Parameter_number=Number of the parameter
               wSubindex_5 : Word;   // Subindex
               wAttribute_NoOfElements_6 : Word := W#16#1000;   // (Attribute=10 Alwais=10)(NoOfParameters=Num of subparameter to Read)
               iParameter_number_6 : Int := 21705;   // Parameter_number=Number of the parameter
               wSubindex_6 : Word;   // Subindex
               wAttribute_NoOfElements_7 : Word := W#16#1000;   // (Attribute=10 Alwais=10)(NoOfParameters=Num of subparameter to Read)
               iParameter_number_7 : Int := 21712;   // Parameter_number=Number of the parameter
               wSubindex_7 : Word;   // Subindex
               wAttribute_NoOfElements_8 : Word := W#16#1000;   // (Attribute=10 Alwais=10)(NoOfParameters=Num of subparameter to Read)
               iParameter_number_8 : Int := 21713;   // Parameter_number=Number of the parameter
               wSubindex_8 : Word;   // Subindex
               wAttribute_NoOfElements_9 : Word := W#16#1000;   // (Attribute=10 Alwais=10)(NoOfParameters=Num of subparameter to Read)
               iParameter_number_9 : Int := 21714;   // Parameter_number=Number of the parameter
               wSubindex_9 : Word;   // Subindex
               wAttribute_NoOfElement_10 : Word := W#16#1000;   // (Attribute=10 Alwais=10)(NoOfParameters=Num of subparameter to Read)
               iParameter_number_10 : Int := 21715;   // Parameter_number=Number of the parameter
               wSubindex_10 : Word;   // Subindex
               wAttribute_NoOfElement_11 : Word := W#16#1000;   // (Attribute=10 Alwais=10)(NoOfParameters=Num of subparameter to Read)
               iParameter_number_11 : Int := 21716;   // Parameter_number=Number of the parameter
               wSubindex_11 : Word;   // Subindex
               wAttribute_NoOfElement_12 : Word := W#16#1000;   // (Attribute=10 Alwais=10)(NoOfParameters=Num of subparameter to Read)
               iParameter_number_12 : Int := 21717;   // Parameter_number=Number of the parameter
               wSubindex_12 : Word;   // Subindex
            END_STRUCT;
            tResponseValues : Struct   // Positive edge record valueas
               wRequest_refere_RequestID : Word;   // (Request_referece=01 Alwais=01 )*(RequestID=01 Read Param)
               wAxis_NoOfParameters : Word;   // (Axis=Num.Object)(NoOfParameters=Num of parameter to Read)
               wFormat_N_Values_1 : Word;   // (Format Parametr) (Number of values)
               dRecordValue_1 : DInt;
               wFormat_N_Values_2 : Word;   // (Format Parametr) (Number of values)
               dRecordValue_2 : DInt;
               wFormat_N_Values_3 : Word;   // (Format Parametr) (Number of values)
               dRecordValue_3 : DInt;
               wFormat_N_Values_4 : Word;   // (Format Parametr) (Number of values)
               dRecordValue_4 : DInt;
               wFormat_N_Values_5 : Word;   // (Format Parametr) (Number of values)
               dRecordValue_5 : DInt;
               wFormat_N_Values_6 : Word;   // (Format Parametr) (Number of values)
               dRecordValue_6 : DInt;
               wFormat_N_Values_7 : Word;   // (Format Parametr) (Number of values)
               dRecordValue_7 : DInt;
               wFormat_N_Values_8 : Word;   // (Format Parametr) (Number of values)
               dRecordValue_8 : DInt;
               wFormat_N_Values_9 : Word;   // (Format Parametr) (Number of values)
               dRecordValue_9 : DInt;
               wFormat_N_Values_10 : Word;   // (Format Parametr) (Number of values)
               dRecordValue_10 : DInt;
               wFormat_N_Values_11 : Word;   // (Format Parametr) (Number of values)
               dRecordValue_11 : DInt;
               wFormat_N_Values_12 : Word;   // (Format Parametr) (Number of values)
               dRecordValue_12 : DInt;
            END_STRUCT;
         END_STRUCT;
      END_STRUCT;
      STC_tW_MngSysReg : Struct   // Managment system register
         tST : Struct